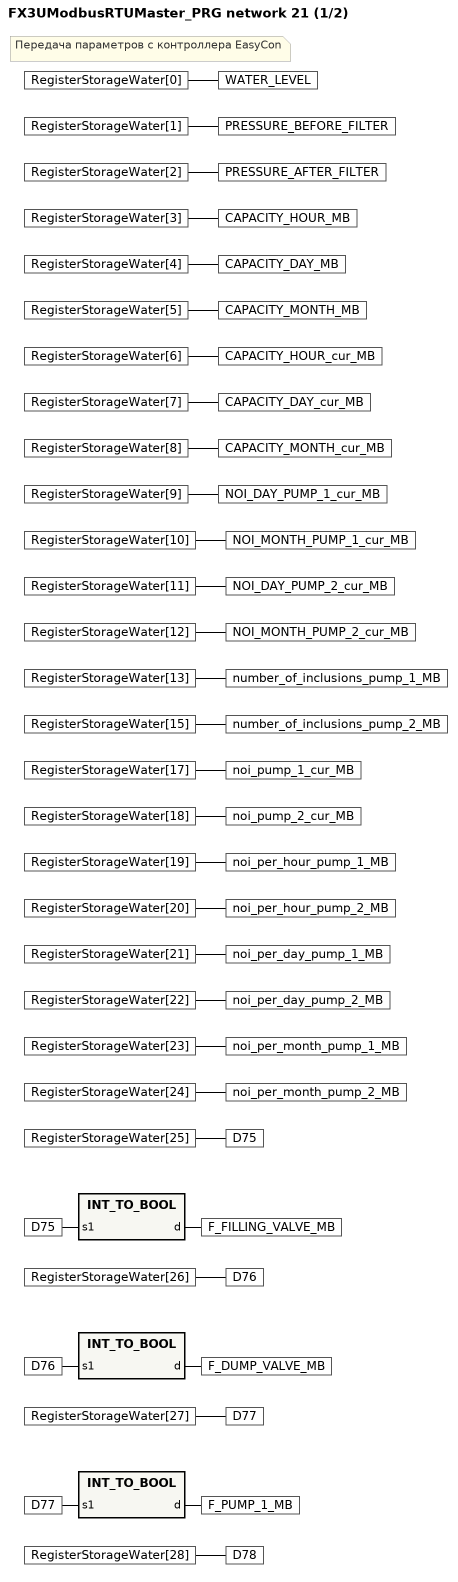
(* [picture p48: structured ladder/FBD of FX3UModbusRTUMaster_PRG, networks 21 to 21] *)
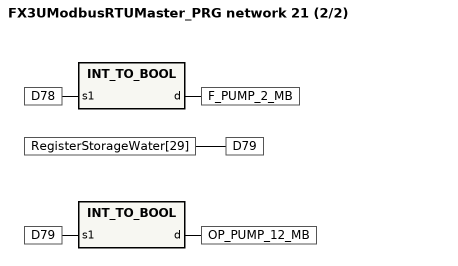
(* network 21 *)
(* Передача параметров с контроллера EasyCon *)
WATER_LEVEL := RegisterStorageWater[0];
PRESSURE_BEFORE_FILTER := RegisterStorageWater[1];
PRESSURE_AFTER_FILTER := RegisterStorageWater[2];
CAPACITY_HOUR_MB := RegisterStorageWater[3];
CAPACITY_DAY_MB := RegisterStorageWater[4];
CAPACITY_MONTH_MB := RegisterStorageWater[5];
CAPACITY_HOUR_cur_MB := RegisterStorageWater[6];
CAPACITY_DAY_cur_MB := RegisterStorageWater[7];
CAPACITY_MONTH_cur_MB := RegisterStorageWater[8];
NOI_DAY_PUMP_1_cur_MB := RegisterStorageWater[9];
NOI_MONTH_PUMP_1_cur_MB := RegisterStorageWater[10];
NOI_DAY_PUMP_2_cur_MB := RegisterStorageWater[11];
NOI_MONTH_PUMP_2_cur_MB := RegisterStorageWater[12];
number_of_inclusions_pump_1_MB := RegisterStorageWater[13];
number_of_inclusions_pump_2_MB := RegisterStorageWater[15];
noi_pump_1_cur_MB := RegisterStorageWater[17];
noi_pump_2_cur_MB := RegisterStorageWater[18];
noi_per_hour_pump_1_MB := RegisterStorageWater[19];
noi_per_hour_pump_2_MB := RegisterStorageWater[20];
noi_per_day_pump_1_MB := RegisterStorageWater[21];
noi_per_day_pump_2_MB := RegisterStorageWater[22];
noi_per_month_pump_1_MB := RegisterStorageWater[23];
noi_per_month_pump_2_MB := RegisterStorageWater[24];
D75 := RegisterStorageWater[25];
F_FILLING_VALVE_MB := INT_TO_BOOL(D75);
D76 := RegisterStorageWater[26];
F_DUMP_VALVE_MB := INT_TO_BOOL(D76);
D77 := RegisterStorageWater[27];
F_PUMP_1_MB := INT_TO_BOOL(D77);
D78 := RegisterStorageWater[28];
F_PUMP_2_MB := INT_TO_BOOL(D78);
D79 := RegisterStorageWater[29];
OP_PUMP_12_MB := INT_TO_BOOL(D79);
END_PROGRAM

PROGRAM VOLTAGE
(* structured ladder/FBD written out as ST: instructions are called as NAME(EN, inputs, outputs); _pN, _eN, _tN stand for wires *)
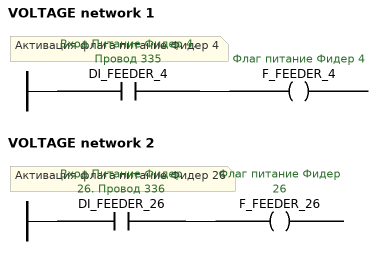
(* network 1 *)
(* Активация флага питание Фидер 4 *)
F_FEEDER_4 := DI_FEEDER_4;
(* network 2 *)
(* Активация флага питание Фидер 26 *)
F_FEEDER_26 := DI_FEEDER_26;
END_PROGRAM
